   END_IF;
   "CV60PosInit" := #_w7;
   IF #_w7 THEN "PLC_to_Epics".CV60.sSetVAuto := 0.0; END_IF;
   #_w8 := #_w2 AND NOT "CV61_ManAuto";
   IF #_w8 THEN
       "unscal_ret_val_7" := UNSCALE(in := 0.0,
                               hi_lim := 100.0,
                               lo_lim := 0.0,
                               bipolar := "always_0",
                               out => "CMD_CV_61");
   END_IF;
   "CV61PosInit" := #_w8;
   IF #_w8 THEN "PLC_to_Epics".CV61.sSetVAuto := 0.0; END_IF;
   IF #_w2 THEN
       "unscal_ret_val_asco_2" := UNSCALE(in := 100.0,
                               hi_lim := 100.0,
                               lo_lim := 0.0,
                               bipolar := "always_0",
                               out => "Sana_ASCO_2");
   END_IF;
   "ASCO2PosInit" := #_w2;
   IF #_w2 THEN
       "ReguleCV61ON" := FALSE;
       "Separators_empty" := FALSE;
   END_IF;
END_REGION

REGION Network 12: Vanne En Position Initial
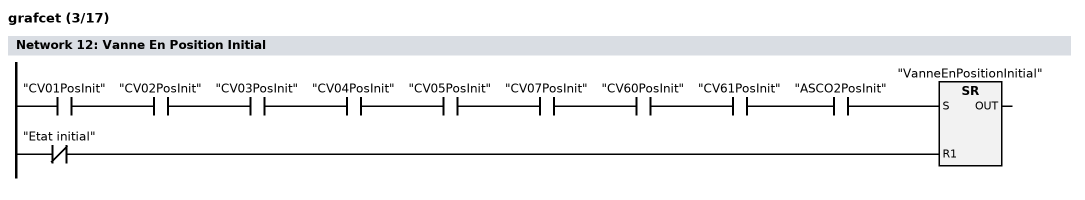
   RUNG wire#powerrail
      Contact( "CV01PosInit" )
      Contact( "CV02PosInit" )
      Contact( "CV03PosInit" )
      Contact( "CV04PosInit" )
      Contact( "CV05PosInit" )
      Contact( "CV07PosInit" )
      Contact( "CV60PosInit" )
      Contact( "CV61PosInit" )
      Contact( "ASCO2PosInit" )
      S_SR(operand := "VanneEnPositionInitial", r1 := wire#w1)
   END_RUNG
   RUNG wire#powerrail
      I_Contact( "Etat initial" )
   END_RUNG wire#w1
   // the same network as SCL:
   IF "CV01PosInit" AND "CV02PosInit" AND "CV03PosInit" AND "CV04PosInit" AND "CV05PosInit" AND "CV07PosInit" AND "CV60PosInit" AND "CV61PosInit" AND "ASCO2PosInit" THEN
       "VanneEnPositionInitial" := TRUE;   // SR flip-flop
   END_IF;
   IF NOT "Etat initial" THEN "VanneEnPositionInitial" := FALSE; END_IF;
END_REGION

REGION Network 13: config vanne etat conditionnement
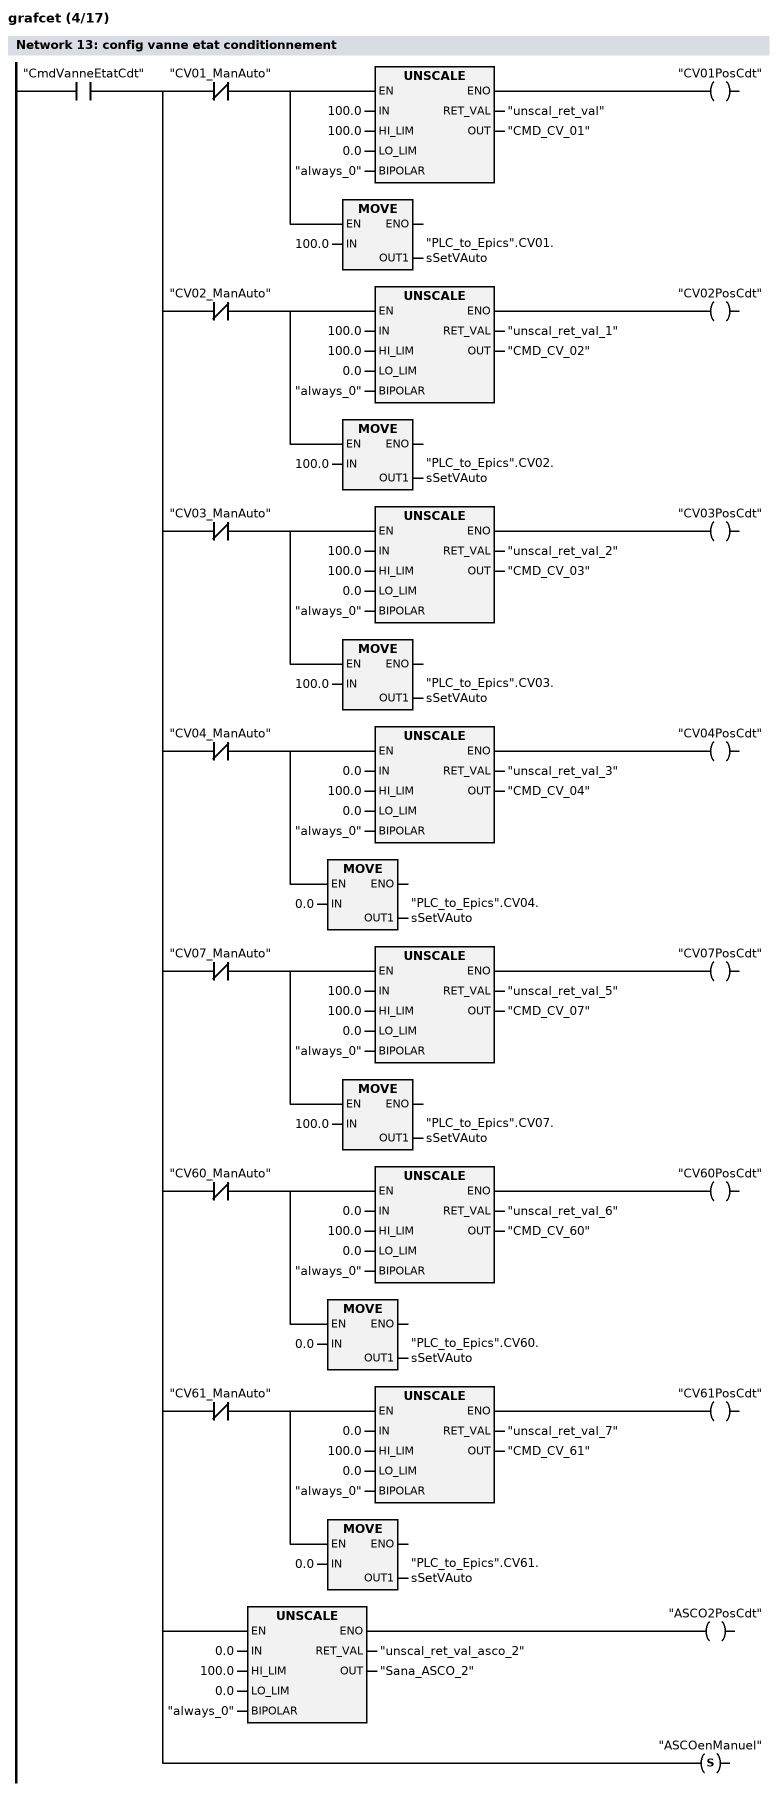
   // ENO of a box is taken as its EN; it also drops when the box reports an error
   #_w1 := "CmdVanneEtatCdt" AND NOT "CV01_ManAuto";
   #_w2 := "CmdVanneEtatCdt";
   IF #_w1 THEN
       "unscal_ret_val" := UNSCALE(IN := 100.0,
                               HI_LIM := 100.0,
                               LO_LIM := 0.0,
                               BIPOLAR := "always_0",
                               OUT => "CMD_CV_01");
   END_IF;
   "CV01PosCdt" := #_w1;
   IF #_w1 THEN "PLC_to_Epics".CV01.sSetVAuto := 100.0; END_IF;
   #_w3 := #_w2 AND NOT "CV02_ManAuto";
   IF #_w3 THEN
       "unscal_ret_val_1" := UNSCALE(IN := 100.0,
                               HI_LIM := 100.0,
                               LO_LIM := 0.0,
                               BIPOLAR := "always_0",
                               OUT => "CMD_CV_02");
   END_IF;
   "CV02PosCdt" := #_w3;
   IF #_w3 THEN "PLC_to_Epics".CV02.sSetVAuto := 100.0; END_IF;
   #_w4 := #_w2 AND NOT "CV03_ManAuto";
   IF #_w4 THEN
       "unscal_ret_val_2" := UNSCALE(IN := 100.0,
                               HI_LIM := 100.0,
                               LO_LIM := 0.0,
                               BIPOLAR := "always_0",
                               OUT => "CMD_CV_03");
   END_IF;
   "CV03PosCdt" := #_w4;
   IF #_w4 THEN "PLC_to_Epics".CV03.sSetVAuto := 100.0; END_IF;
   #_w5 := #_w2 AND NOT "CV04_ManAuto";
   IF #_w5 THEN
       "unscal_ret_val_3" := UNSCALE(IN := 0.0,
                               HI_LIM := 100.0,
                               LO_LIM := 0.0,
                               BIPOLAR := "always_0",
                               OUT => "CMD_CV_04");
   END_IF;
   "CV04PosCdt" := #_w5;
   IF #_w5 THEN "PLC_to_Epics".CV04.sSetVAuto := 0.0; END_IF;
   #_w6 := #_w2 AND NOT "CV07_ManAuto";
   IF #_w6 THEN
       "unscal_ret_val_5" := UNSCALE(IN := 100.0,
                               HI_LIM := 100.0,
                               LO_LIM := 0.0,
                               BIPOLAR := "always_0",
                               OUT => "CMD_CV_07");
   END_IF;
   "CV07PosCdt" := #_w6;
   IF #_w6 THEN "PLC_to_Epics".CV07.sSetVAuto := 100.0; END_IF;
   #_w7 := #_w2 AND NOT "CV60_ManAuto";
   IF #_w7 THEN
       "unscal_ret_val_6" := UNSCALE(IN := 0.0,
                               HI_LIM := 100.0,
                               LO_LIM := 0.0,
                               BIPOLAR := "always_0",
                               OUT => "CMD_CV_60");
   END_IF;
   "CV60PosCdt" := #_w7;
   IF #_w7 THEN "PLC_to_Epics".CV60.sSetVAuto := 0.0; END_IF;
   #_w8 := #_w2 AND NOT "CV61_ManAuto";
   IF #_w8 THEN
       "unscal_ret_val_7" := UNSCALE(IN := 0.0,
                               HI_LIM := 100.0,
                               LO_LIM := 0.0,
                               BIPOLAR := "always_0",
                               OUT => "CMD_CV_61");
   END_IF;
   "CV61PosCdt" := #_w8;
   IF #_w8 THEN "PLC_to_Epics".CV61.sSetVAuto := 0.0; END_IF;
   IF #_w2 THEN
       "unscal_ret_val_asco_2" := UNSCALE(IN := 0.0,
                               HI_LIM := 100.0,
                               LO_LIM := 0.0,
                               BIPOLAR := "always_0",
                               OUT => "Sana_ASCO_2");
   END_IF;
   "ASCO2PosCdt" := #_w2;
   IF #_w2 THEN "ASCOenManuel" := TRUE; END_IF;
END_REGION

REGION Network 14: Vanne En Position Cdt
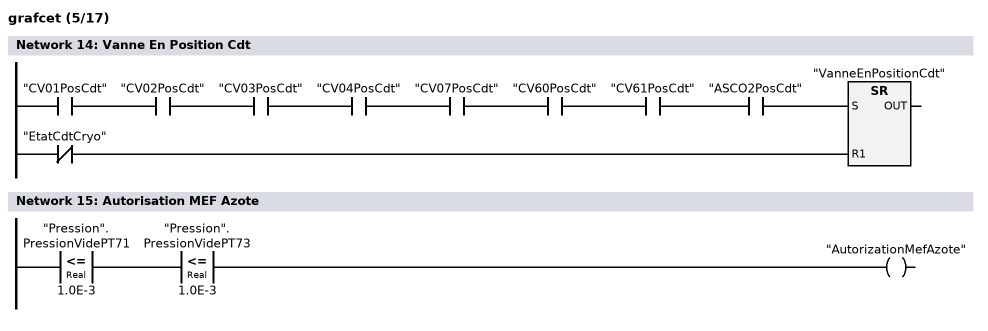
   RUNG wire#powerrail
      Contact( "CV01PosCdt" )
      Contact( "CV02PosCdt" )
      Contact( "CV03PosCdt" )
      Contact( "CV04PosCdt" )
      Contact( "CV07PosCdt" )
      Contact( "CV60PosCdt" )
      Contact( "CV61PosCdt" )
      Contact( "ASCO2PosCdt" )
      S_SR(operand := "VanneEnPositionCdt", r1 := wire#w1)
   END_RUNG
   RUNG wire#powerrail
      I_Contact( "EtatCdtCryo" )
   END_RUNG wire#w1
   // the same network as SCL:
   IF "CV01PosCdt" AND "CV02PosCdt" AND "CV03PosCdt" AND "CV04PosCdt" AND "CV07PosCdt" AND "CV60PosCdt" AND "CV61PosCdt" AND "ASCO2PosCdt" THEN
       "VanneEnPositionCdt" := TRUE;   // SR flip-flop
   END_IF;
   IF NOT "EtatCdtCryo" THEN "VanneEnPositionCdt" := FALSE; END_IF;
END_REGION

REGION Network 15: Autorisation MEF Azote
   RUNG wire#powerrail
      { S7_Templates := "SrcType := Real" } LE_Contact(in1 := "Pression".PressionVidePT71, in2 := 1.0E-3)
      { S7_Templates := "SrcType := Real" } LE_Contact(in1 := "Pression".PressionVidePT73, in2 := 1.0E-3)
      Coil( "AutorizationMefAzote" )
   END_RUNG
   // the same network as SCL:
   "AutorizationMefAzote" := ("Pression".PressionVidePT71 <= 1.0E-3) AND ("Pression".PressionVidePT73 <= 1.0E-3);
END_REGION

REGION Network 16: config vannes init mode & regule cv61 on
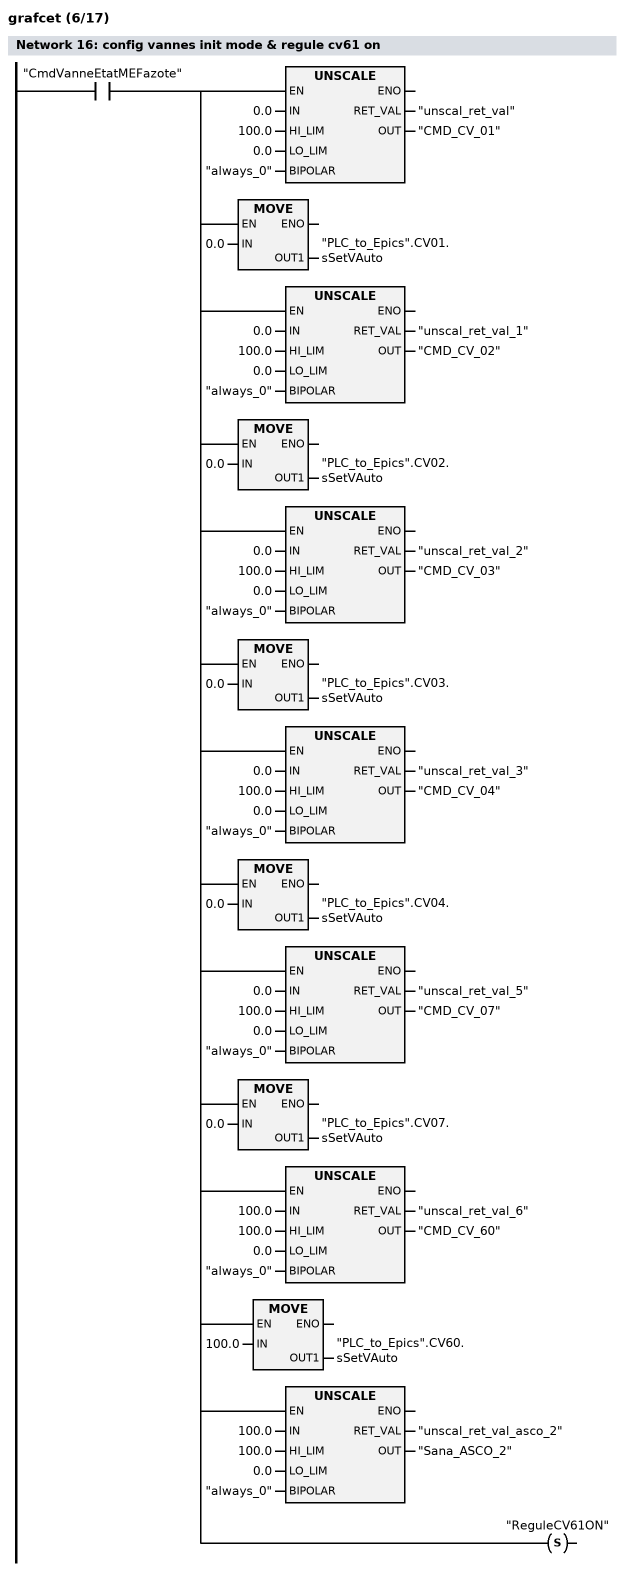
   #_w1 := "CmdVanneEtatMEFazote";
   IF #_w1 THEN
       "unscal_ret_val" := UNSCALE(in := 0.0,
                               hi_lim := 100.0,
                               lo_lim := 0.0,
                               bipolar := "always_0",
                               out => "CMD_CV_01");
       "PLC_to_Epics".CV01.sSetVAuto := 0.0;
       "unscal_ret_val_1" := UNSCALE(in := 0.0,
                               hi_lim := 100.0,
                               lo_lim := 0.0,
                               bipolar := "always_0",
                               out => "CMD_CV_02");
       "PLC_to_Epics".CV02.sSetVAuto := 0.0;
       "unscal_ret_val_2" := UNSCALE(in := 0.0,
                               hi_lim := 100.0,
                               lo_lim := 0.0,
                               bipolar := "always_0",
                               out => "CMD_CV_03");
       "PLC_to_Epics".CV03.sSetVAuto := 0.0;
       "unscal_ret_val_3" := UNSCALE(in := 0.0,
                               hi_lim := 100.0,
                               lo_lim := 0.0,
                               bipolar := "always_0",
                               out => "CMD_CV_04");
       "PLC_to_Epics".CV04.sSetVAuto := 0.0;
       "unscal_ret_val_5" := UNSCALE(in := 0.0,
                               hi_lim := 100.0,
                               lo_lim := 0.0,
                               bipolar := "always_0",
                               out => "CMD_CV_07");
       "PLC_to_Epics".CV07.sSetVAuto := 0.0;
       "unscal_ret_val_6" := UNSCALE(in := 100.0,
                               hi_lim := 100.0,
                               lo_lim := 0.0,
                               bipolar := "always_0",
                               out => "CMD_CV_60");
       "PLC_to_Epics".CV60.sSetVAuto := 100.0;
       "unscal_ret_val_asco_2" := UNSCALE(in := 100.0,
                               hi_lim := 100.0,
                               lo_lim := 0.0,
                               bipolar := "always_0",
                               out => "Sana_ASCO_2");
       "ReguleCV61ON" := TRUE;
   END_IF;
END_REGION

REGION Network 17: Régule CV61 seuil (desactive)
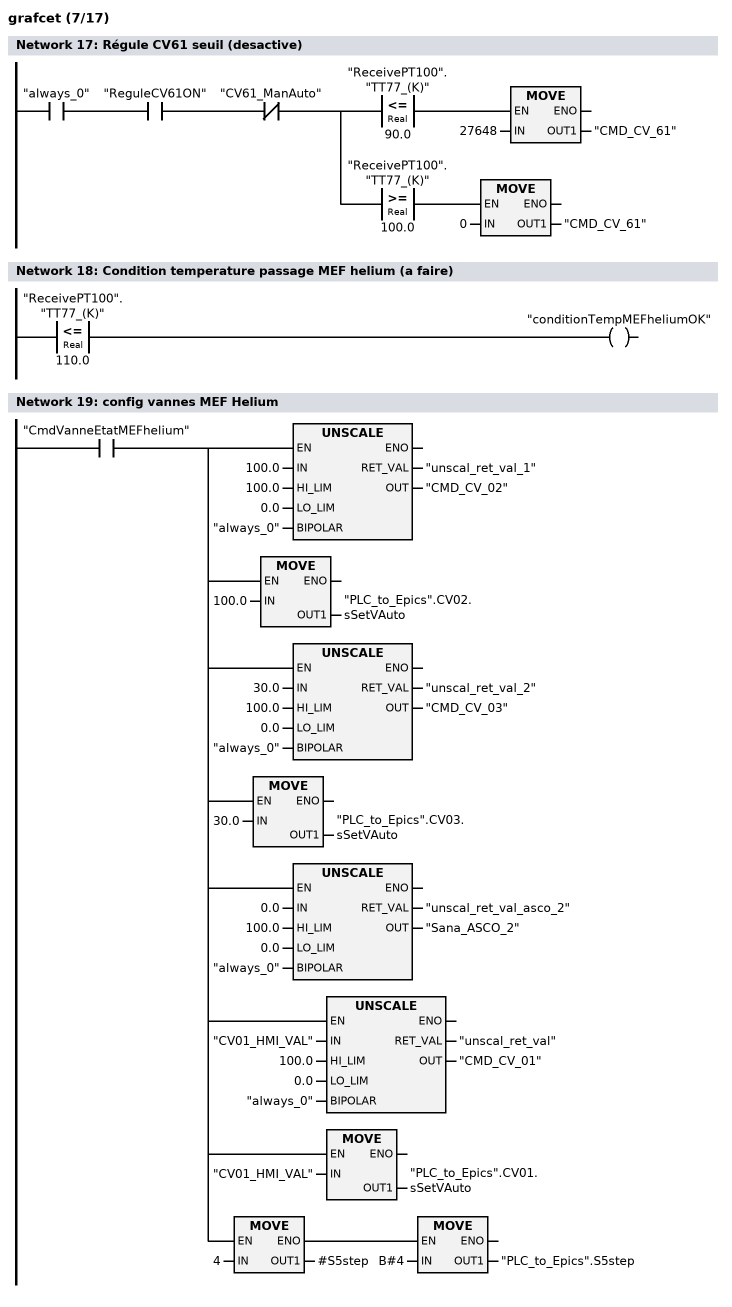
   RUNG wire#powerrail
      Contact( "always_0" )
      Contact( "ReguleCV61ON" )
      I_Contact( "CV61_ManAuto" )
      wire#w1
      { S7_Templates := "SrcType := Real" } LE_Contact(in1 := "ReceivePT100"."TT77_(K)", in2 := 90.0)
      { S7_GenerateENO := "TRUE" } Move(in := 27648, out1 => "CMD_CV_61")
   END_RUNG
   RUNG wire#w1
      { S7_Templates := "SrcType := Real" } GE_Contact(in1 := "ReceivePT100"."TT77_(K)", in2 := 100.0)
      { S7_GenerateENO := "TRUE" } Move(in := 0, out1 => "CMD_CV_61")
   END_RUNG
   // the same network as SCL:
   #_w1 := "always_0" AND "ReguleCV61ON" AND NOT "CV61_ManAuto";
   IF #_w1 AND ("ReceivePT100"."TT77_(K)" <= 90.0) THEN "CMD_CV_61" := 27648; END_IF;
   IF #_w1 AND ("ReceivePT100"."TT77_(K)" >= 100.0) THEN "CMD_CV_61" := 0; END_IF;
END_REGION

REGION Network 18: Condition temperature passage MEF helium (a faire)
   RUNG wire#powerrail
      { S7_Templates := "SrcType := Real" } LE_Contact(in1 := "ReceivePT100"."TT77_(K)", in2 := 110.0)
      Coil( "conditionTempMEFheliumOK" )
   END_RUNG
   // the same network as SCL:
   "conditionTempMEFheliumOK" := "ReceivePT100"."TT77_(K)" <= 110.0;
END_REGION

REGION Network 19: config vannes MEF Helium
   // ENO of a box is taken as its EN; it also drops when the box reports an error
   #_w1 := "CmdVanneEtatMEFhelium";
   IF #_w1 THEN
       "unscal_ret_val_1" := UNSCALE(IN := 100.0,
                               HI_LIM := 100.0,
                               LO_LIM := 0.0,
                               BIPOLAR := "always_0",
                               OUT => "CMD_CV_02");
       "PLC_to_Epics".CV02.sSetVAuto := 100.0;
       "unscal_ret_val_2" := UNSCALE(IN := 30.0,
                               HI_LIM := 100.0,
                               LO_LIM := 0.0,
                               BIPOLAR := "always_0",
                               OUT => "CMD_CV_03");
       "PLC_to_Epics".CV03.sSetVAuto := 30.0;
       "unscal_ret_val_asco_2" := UNSCALE(IN := 0.0,
                               HI_LIM := 100.0,
                               LO_LIM := 0.0,
                               BIPOLAR := "always_0",
                               OUT => "Sana_ASCO_2");
       "unscal_ret_val" := UNSCALE(IN := "CV01_HMI_VAL",
                               HI_LIM := 100.0,
                               LO_LIM := 0.0,
                               BIPOLAR := "always_0",
                               OUT => "CMD_CV_01");
       "PLC_to_Epics".CV01.sSetVAuto := "CV01_HMI_VAL";
       #S5step := 4;
       "PLC_to_Epics".S5step := B#4;
   END_IF;
END_REGION

REGION Network 20: LHe cooling down - Set step 6 (maybe setting CV03 is not needed here (done in the next network)!!!!!
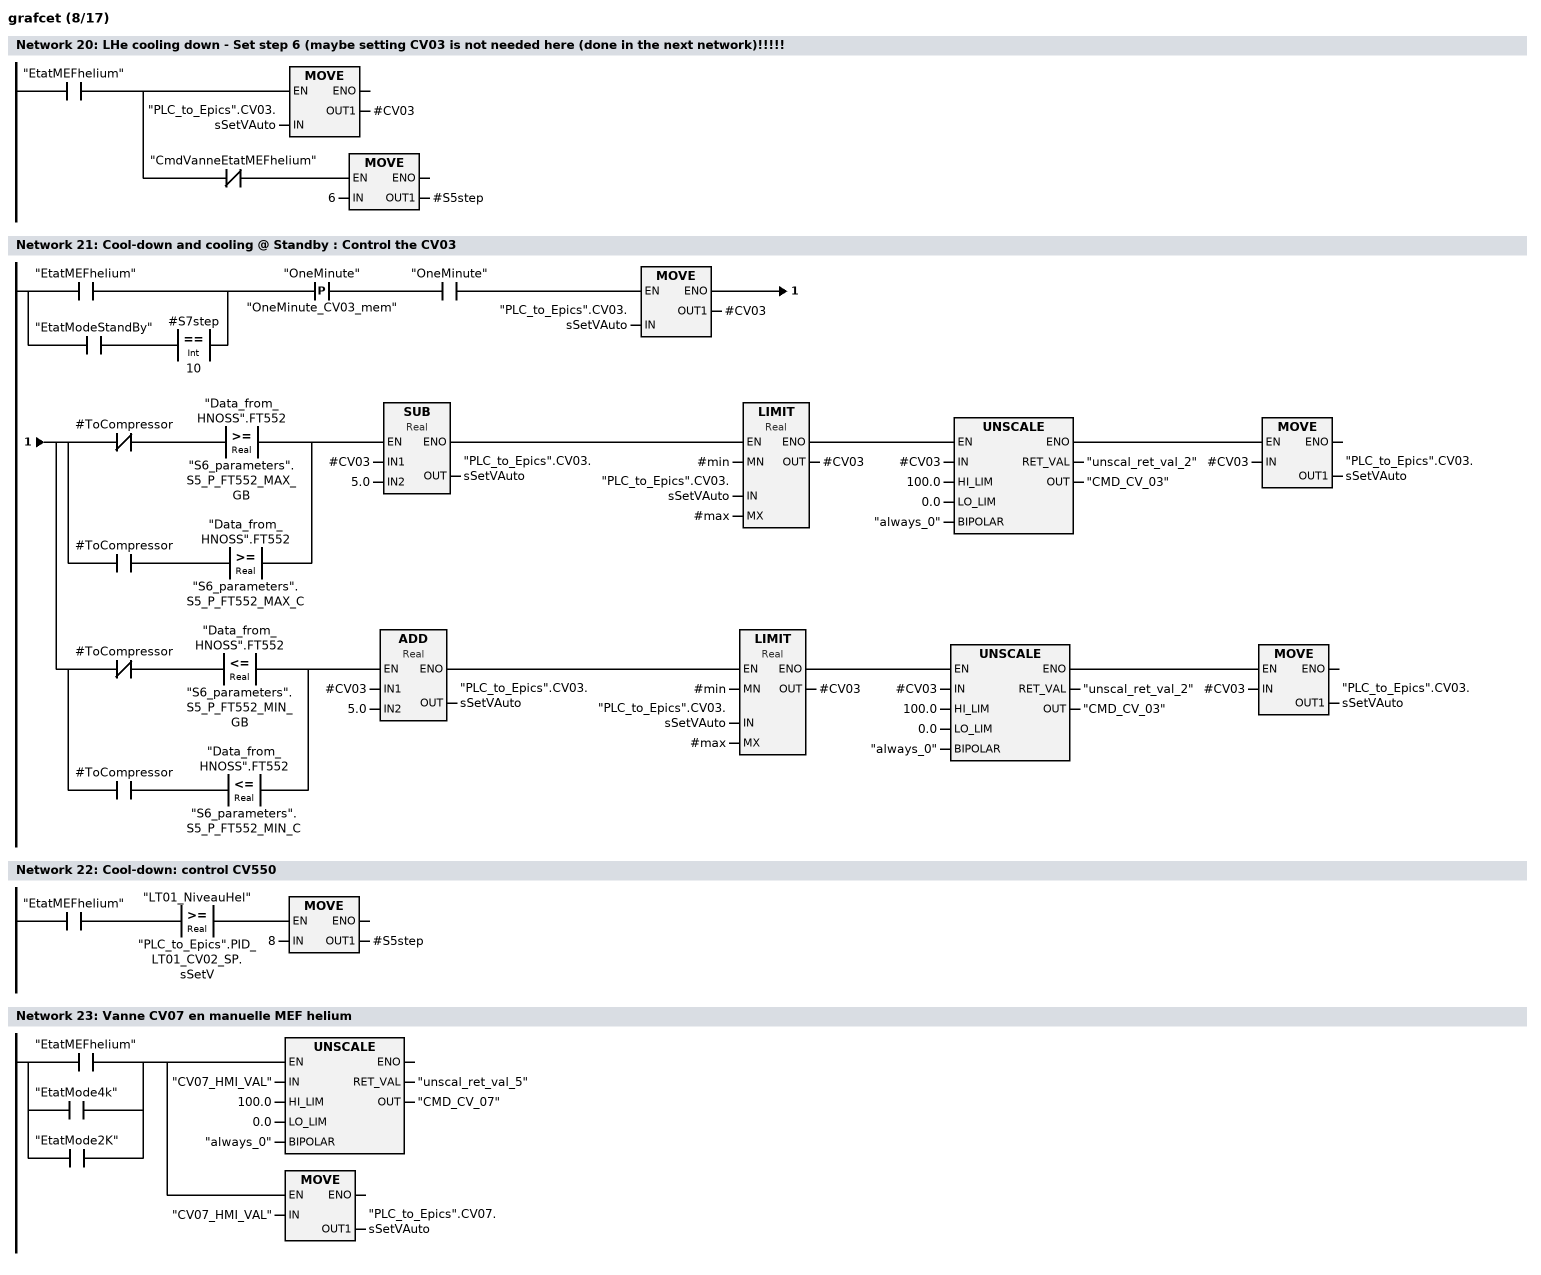
   RUNG wire#powerrail
      Contact( "EtatMEFhelium" )
      wire#w1
      { S7_GenerateENO := "TRUE" } Move(in := "PLC_to_Epics".CV03.sSetVAuto, out1 => #CV03)
   END_RUNG
   RUNG wire#w1
      I_Contact( "CmdVanneEtatMEFhelium" )
      { S7_GenerateENO := "TRUE" } Move(in := 6, out1 => #S5step)
   END_RUNG
   // the same network as SCL:
   IF "EtatMEFhelium" THEN #CV03 := "PLC_to_Epics".CV03.sSetVAuto; END_IF;
   IF "EtatMEFhelium" AND NOT "CmdVanneEtatMEFhelium" THEN #S5step := 6; END_IF;
END_REGION

REGION Network 21: Cool-down and cooling @ Standby : Control the CV03
   // ENO of a box is taken as its EN; it also drops when the box reports an error
   #_w1 := ("EtatMEFhelium" OR ("EtatModeStandBy" AND (#S7step = 10))) AND "OneMinute" AND NOT "OneMinute_CV03_mem";   // rising edge of "OneMinute"
   "OneMinute_CV03_mem" := "OneMinute";
   #_w2 := #_w1 AND "OneMinute";
   IF #_w2 THEN #CV03 := "PLC_to_Epics".CV03.sSetVAuto; END_IF;
   IF #_w2 AND ((NOT #ToCompressor AND ("Data_from_HNOSS".FT552 >= "S6_parameters".S5_P_FT552_MAX_GB)) OR (#ToCompressor AND ("Data_from_HNOSS".FT552 >= "S6_parameters".S5_P_FT552_MAX_C))) THEN
       "PLC_to_Epics".CV03.sSetVAuto := #CV03 - 5.0;
       #CV03 := LIMIT(MN := #min, IN := "PLC_to_Epics".CV03.sSetVAuto, MX := #max);
   END_IF;
   #_w3 := #_w2 AND ((NOT #ToCompressor AND ("Data_from_HNOSS".FT552 >= "S6_parameters".S5_P_FT552_MAX_GB)) OR (#ToCompressor AND ("Data_from_HNOSS".FT552 >= "S6_parameters".S5_P_FT552_MAX_C)));
   IF #_w3 THEN
       "unscal_ret_val_2" := UNSCALE(IN := #CV03,
                               HI_LIM := 100.0,
                               LO_LIM := 0.0,
                               BIPOLAR := "always_0",
                               OUT => "CMD_CV_03");
       "PLC_to_Epics".CV03.sSetVAuto := #CV03;
   END_IF;
   IF #_w2 AND ((NOT #ToCompressor AND ("Data_from_HNOSS".FT552 <= "S6_parameters".S5_P_FT552_MIN_GB)) OR (#ToCompressor AND ("Data_from_HNOSS".FT552 <= "S6_parameters".S5_P_FT552_MIN_C))) THEN
       "PLC_to_Epics".CV03.sSetVAuto := #CV03 + 5.0;
       #CV03 := LIMIT(MN := #min, IN := "PLC_to_Epics".CV03.sSetVAuto, MX := #max);
   END_IF;
   #_w4 := #_w2 AND ((NOT #ToCompressor AND ("Data_from_HNOSS".FT552 <= "S6_parameters".S5_P_FT552_MIN_GB)) OR (#ToCompressor AND ("Data_from_HNOSS".FT552 <= "S6_parameters".S5_P_FT552_MIN_C)));
   IF #_w4 THEN
       "unscal_ret_val_2" := UNSCALE(IN := #CV03,
                               HI_LIM := 100.0,
                               LO_LIM := 0.0,
                               BIPOLAR := "always_0",
                               OUT => "CMD_CV_03");
       "PLC_to_Epics".CV03.sSetVAuto := #CV03;
   END_IF;
END_REGION

REGION Network 22: Cool-down: control CV550
   RUNG wire#powerrail
      Contact( "EtatMEFhelium" )
      { S7_Templates := "SrcType := Real" } GE_Contact(in1 := "LT01_NiveauHel", in2 := "PLC_to_Epics".PID_LT01_CV02_SP.sSetV)
      { S7_GenerateENO := "TRUE" } Move(in := 8, out1 => #S5step)
   END_RUNG
   // the same network as SCL:
   IF "EtatMEFhelium" AND ("LT01_NiveauHel" >= "PLC_to_Epics".PID_LT01_CV02_SP.sSetV) THEN
       #S5step := 8;
   END_IF;
END_REGION

REGION Network 23: Vanne CV07 en manuelle MEF helium
   #_w1 := "EtatMEFhelium" OR "EtatMode4k" OR "EtatMode2K";
   IF #_w1 THEN
       "unscal_ret_val_5" := UNSCALE(in := "CV07_HMI_VAL",
                               hi_lim := 100.0,
                               lo_lim := 0.0,
                               bipolar := "always_0",
                               out => "CMD_CV_07");
       "PLC_to_Epics".CV07.sSetVAuto := "CV07_HMI_VAL";
   END_IF;
END_REGION

REGION Network 24: Vanne CV01 en manuelle MEF helium
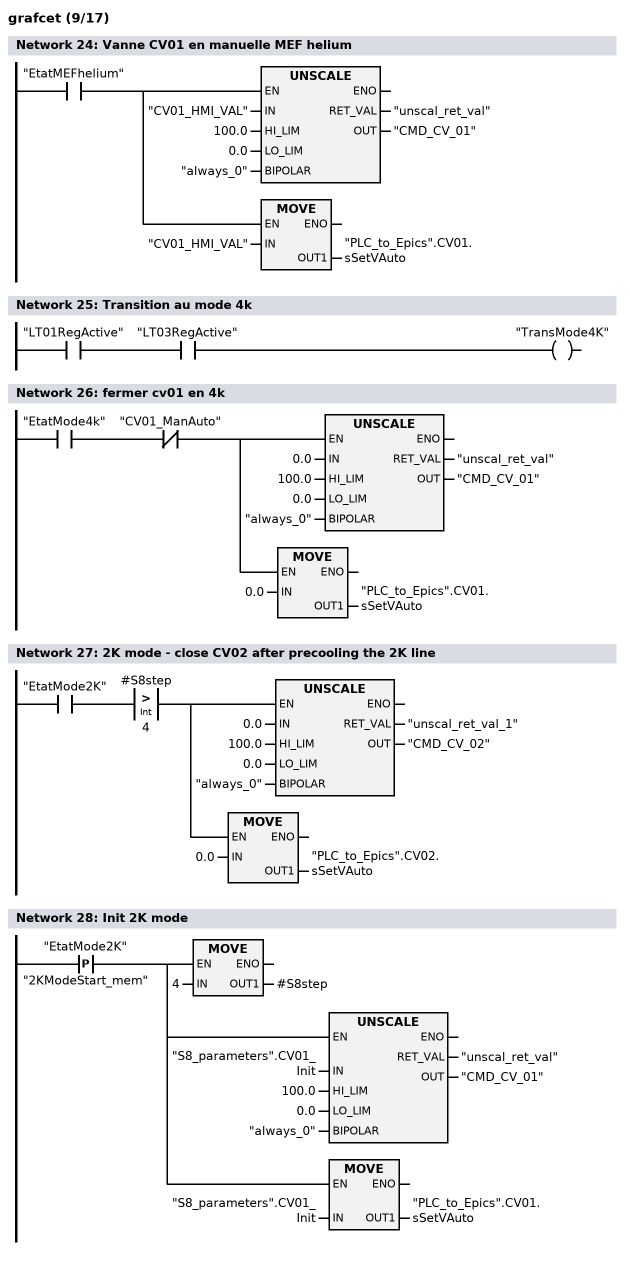
   #_w1 := "EtatMEFhelium";
   IF #_w1 THEN
       "unscal_ret_val" := UNSCALE(in := "CV01_HMI_VAL",
                               hi_lim := 100.0,
                               lo_lim := 0.0,
                               bipolar := "always_0",
                               out => "CMD_CV_01");
       "PLC_to_Epics".CV01.sSetVAuto := "CV01_HMI_VAL";
   END_IF;
END_REGION

REGION Network 25: Transition au mode 4k
   RUNG wire#powerrail
      Contact( "LT01RegActive" )
      Contact( "LT03RegActive" )
      Coil( "TransMode4K" )
   END_RUNG
   // the same network as SCL:
   "TransMode4K" := "LT01RegActive" AND "LT03RegActive";
END_REGION

REGION Network 26: fermer cv01 en 4k
   #_w1 := "EtatMode4k" AND NOT "CV01_ManAuto";
   IF #_w1 THEN
       "unscal_ret_val" := UNSCALE(in := 0.0,
                               hi_lim := 100.0,
                               lo_lim := 0.0,
                               bipolar := "always_0",
                               out => "CMD_CV_01");
       "PLC_to_Epics".CV01.sSetVAuto := 0.0;
   END_IF;
END_REGION

REGION Network 27: 2K mode - close CV02 after precooling the 2K line
   #_w1 := "EtatMode2K" AND (#S8step > 4);
   IF #_w1 THEN
       "unscal_ret_val_1" := UNSCALE(IN := 0.0,
                               HI_LIM := 100.0,
                               LO_LIM := 0.0,
                               BIPOLAR := "always_0",
                               OUT => "CMD_CV_02");
       "PLC_to_Epics".CV02.sSetVAuto := 0.0;
   END_IF;
END_REGION

REGION Network 28: Init 2K mode
   #_w1 := "EtatMode2K" AND NOT "2KModeStart_mem";   // rising edge of "EtatMode2K"
   "2KModeStart_mem" := "EtatMode2K";
   IF #_w1 THEN
       #S8step := 4;
       "unscal_ret_val" := UNSCALE(IN := "S8_parameters".CV01_Init,
                               HI_LIM := 100.0,
                               LO_LIM := 0.0,
                               BIPOLAR := "always_0",
                               OUT => "CMD_CV_01");
       "PLC_to_Epics".CV01.sSetVAuto := "S8_parameters".CV01_Init;
   END_IF;
END_REGION

REGION Network 29: 2K mode - precooling (step4)
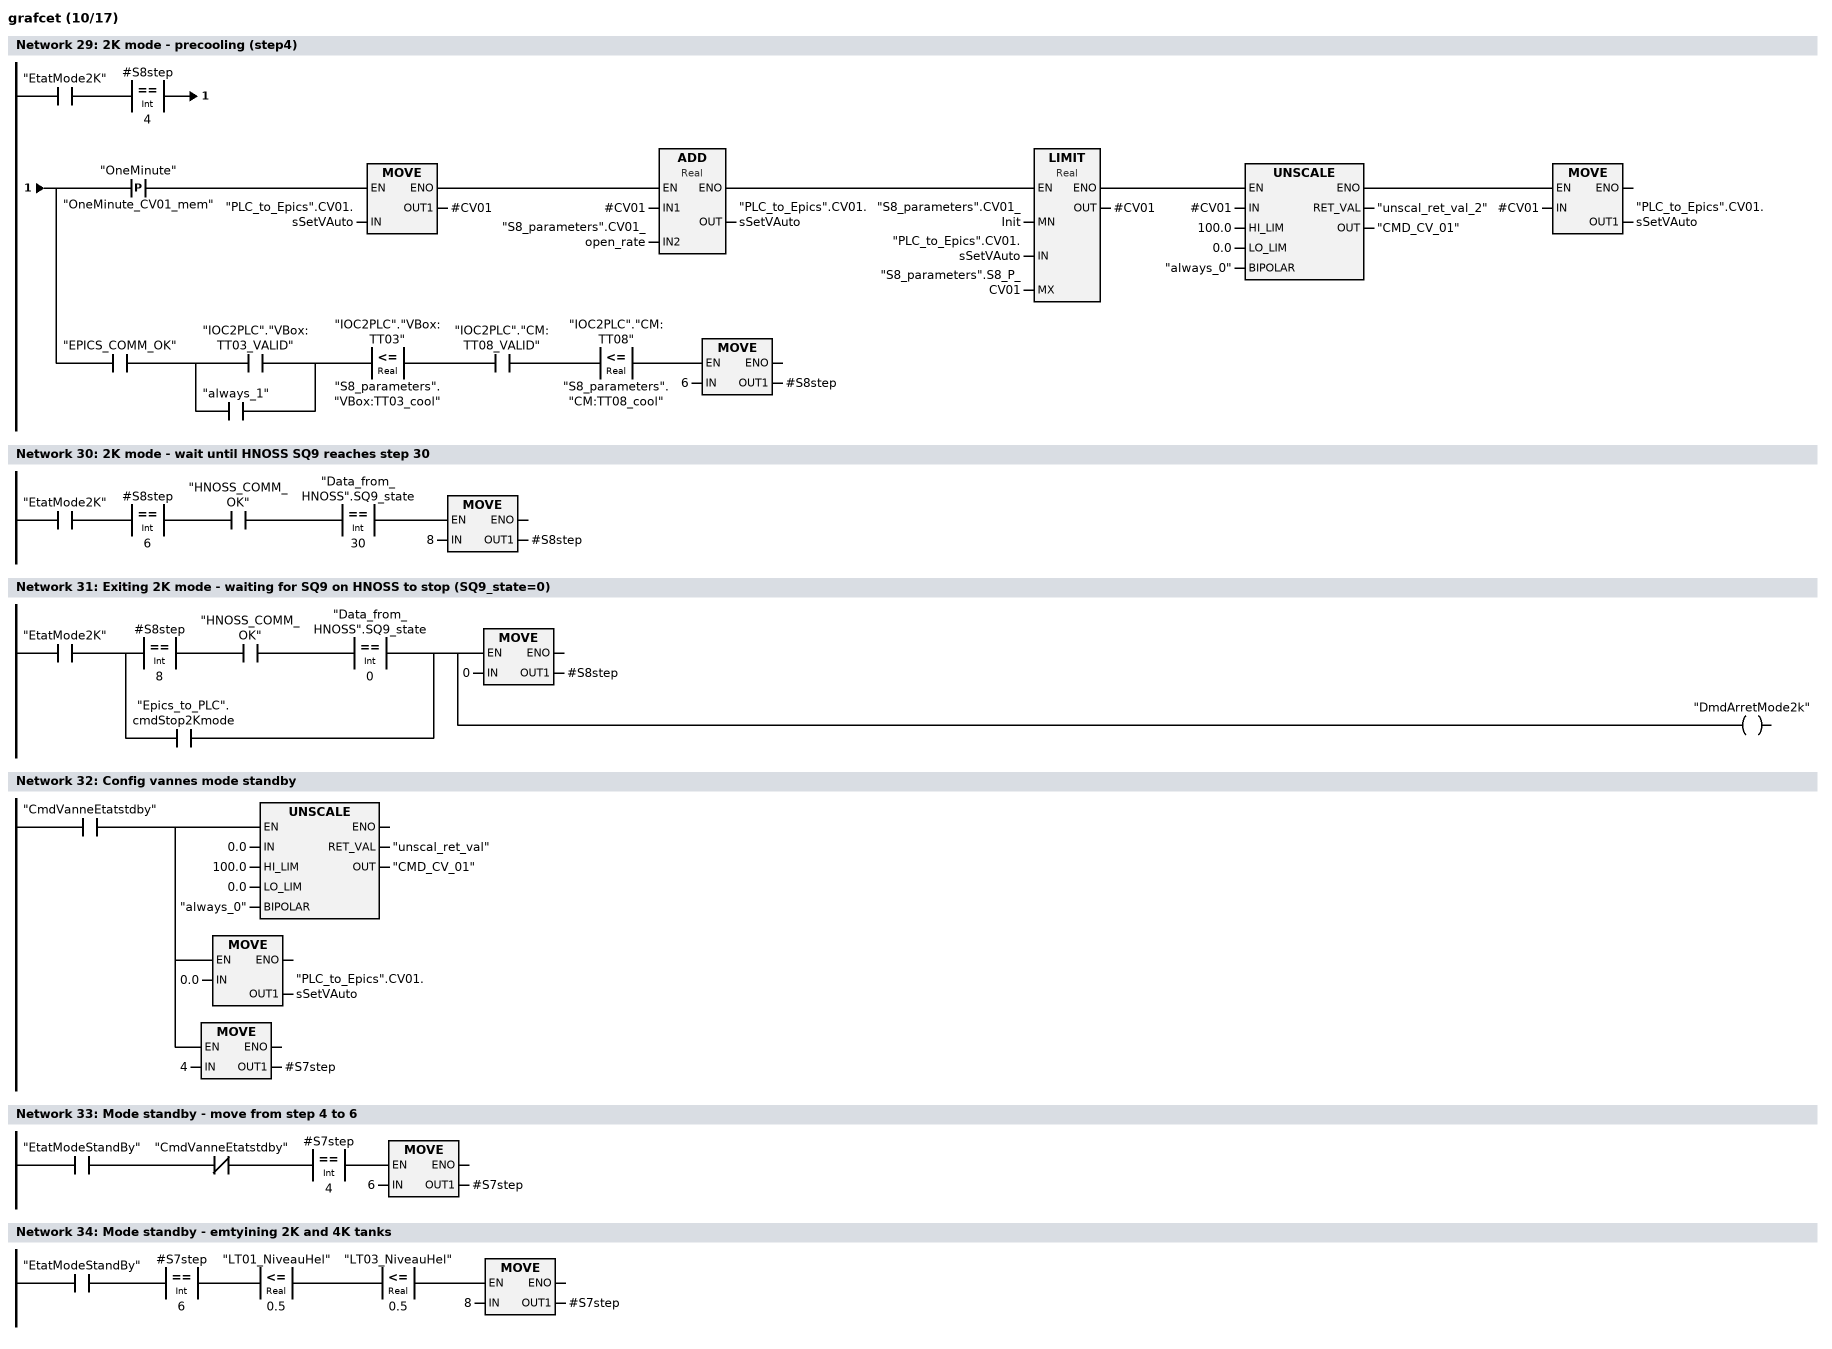
   // ENO of a box is taken as its EN; it also drops when the box reports an error
   #_w1 := "EtatMode2K" AND (#S8step = 4);
   #_w2 := #_w1 AND "OneMinute" AND NOT "OneMinute_CV01_mem";   // rising edge of "OneMinute"
   "OneMinute_CV01_mem" := "OneMinute";
   IF #_w2 THEN
       #CV01 := "PLC_to_Epics".CV01.sSetVAuto;
       "PLC_to_Epics".CV01.sSetVAuto := #CV01 + "S8_parameters".CV01_open_rate;
       #CV01 := LIMIT(MN := "S8_parameters".CV01_Init, IN := "PLC_to_Epics".CV01.sSetVAuto, MX := "S8_parameters".S8_P_CV01);
       "unscal_ret_val_2" := UNSCALE(IN := #CV01,
                               HI_LIM := 100.0,
                               LO_LIM := 0.0,
                               BIPOLAR := "always_0",
                               OUT => "CMD_CV_01");
       "PLC_to_Epics".CV01.sSetVAuto := #CV01;
   END_IF;
   IF #_w1 AND "EPICS_COMM_OK" AND ("IOC2PLC"."VBox:TT03_VALID" OR "always_1") AND ("IOC2PLC"."VBox:TT03" <= "S8_parameters"."VBox:TT03_cool") AND "IOC2PLC"."CM:TT08_VALID" AND ("IOC2PLC"."CM:TT08" <= "S8_parameters"."CM:TT08_cool") THEN
       #S8step := 6;
   END_IF;
END_REGION

REGION Network 30: 2K mode - wait until HNOSS SQ9 reaches step 30
   RUNG wire#powerrail
      Contact( "EtatMode2K" )
      { S7_Templates := "SrcType := Int" } EQ_Contact(in1 := #S8step, in2 := 6)
      Contact( "HNOSS_COMM_OK" )
      { S7_Templates := "SrcType := Int" } EQ_Contact(in1 := "Data_from_HNOSS".SQ9_state, in2 := 30)
      { S7_GenerateENO := "TRUE" } Move(in := 8, out1 => #S8step)
   END_RUNG
   // the same network as SCL:
   IF "EtatMode2K" AND (#S8step = 6) AND "HNOSS_COMM_OK" AND ("Data_from_HNOSS".SQ9_state = 30) THEN
       #S8step := 8;
   END_IF;
END_REGION

REGION Network 31: Exiting 2K mode - waiting for SQ9 on HNOSS to stop (SQ9_state=0)
   RUNG wire#powerrail
      Contact( "EtatMode2K" )
      wire#w1
      { S7_Templates := "SrcType := Int" } EQ_Contact(in1 := #S8step, in2 := 8)
      Contact( "HNOSS_COMM_OK" )
      { S7_Templates := "SrcType := Int" } EQ_Contact(in1 := "Data_from_HNOSS".SQ9_state, in2 := 0)
      wire#w2
      { S7_GenerateENO := "TRUE" } Move(in := 0, out1 => #S8step)
   END_RUNG
   RUNG wire#w1
      Contact( "Epics_to_PLC".cmdStop2Kmode )
   END_RUNG wire#w2
   RUNG wire#w2
      Coil( "DmdArretMode2k" )
   END_RUNG
   // the same network as SCL:
   #_w1 := "EtatMode2K" AND (((#S8step = 8) AND "HNOSS_COMM_OK" AND ("Data_from_HNOSS".SQ9_state = 0)) OR "Epics_to_PLC".cmdStop2Kmode);
   IF #_w1 THEN #S8step := 0; END_IF;
   "DmdArretMode2k" := #_w1;
END_REGION

REGION Network 32: Config vannes mode standby
   #_w1 := "CmdVanneEtatstdby";
   IF #_w1 THEN
       "unscal_ret_val" := UNSCALE(IN := 0.0,
                               HI_LIM := 100.0,
                               LO_LIM := 0.0,
                               BIPOLAR := "always_0",
                               OUT => "CMD_CV_01");
       "PLC_to_Epics".CV01.sSetVAuto := 0.0;
       #S7step := 4;
   END_IF;
END_REGION

REGION Network 33: Mode standby - move from step 4 to 6
   RUNG wire#powerrail
      Contact( "EtatModeStandBy" )
      I_Contact( "CmdVanneEtatstdby" )
      { S7_Templates := "SrcType := Int" } EQ_Contact(in1 := #S7step, in2 := 4)
      { S7_GenerateENO := "TRUE" } Move(in := 6, out1 => #S7step)
   END_RUNG
   // the same network as SCL:
   IF "EtatModeStandBy" AND NOT "CmdVanneEtatstdby" AND (#S7step = 4) THEN #S7step := 6; END_IF;
END_REGION

REGION Network 34: Mode standby - emtyining 2K and 4K tanks
   RUNG wire#powerrail
      Contact( "EtatModeStandBy" )
      { S7_Templates := "SrcType := Int" } EQ_Contact(in1 := #S7step, in2 := 6)
      { S7_Templates := "SrcType := Real" } LE_Contact(in1 := "LT01_NiveauHel", in2 := 0.5)
      { S7_Templates := "SrcType := Real" } LE_Contact(in1 := "LT03_NiveauHel", in2 := 0.5)
      { S7_GenerateENO := "TRUE" } Move(in := 8, out1 => #S7step)
   END_RUNG
   // the same network as SCL:
   IF "EtatModeStandBy" AND (#S7step = 6) AND ("LT01_NiveauHel" <= 0.5) AND ("LT03_NiveauHel" <= 0.5) THEN
       #S7step := 8;
   END_IF;
END_REGION

REGION Network 35: Mode standby - warming up (step8) and cooling (step10)
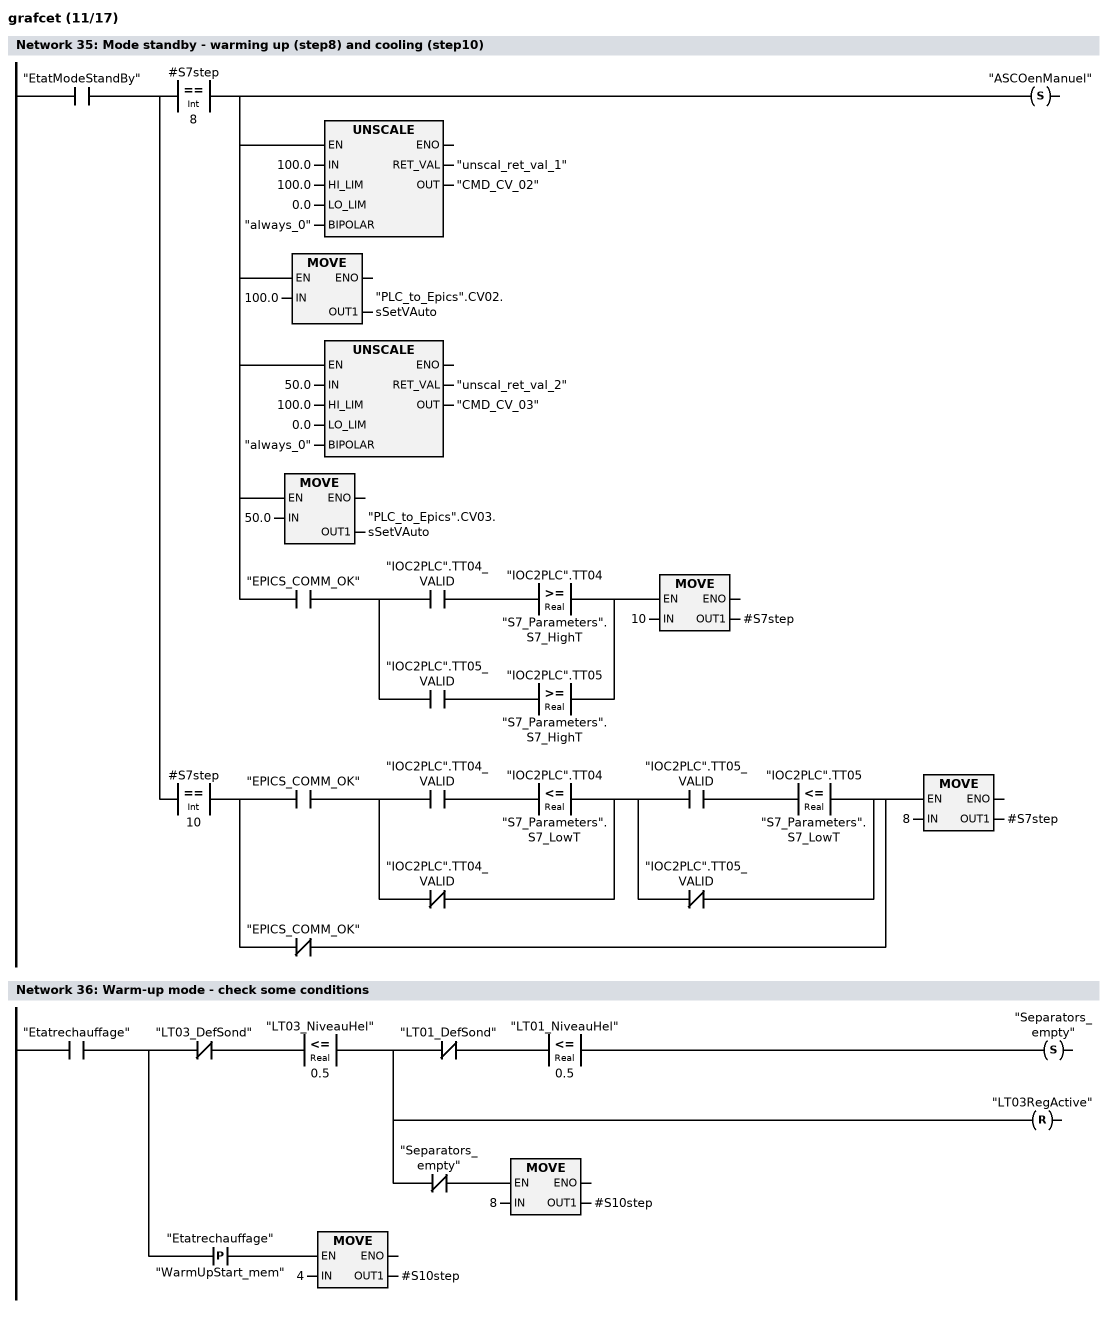
   #_w1 := "EtatModeStandBy" AND (#S7step = 8);
   IF #_w1 THEN "ASCOenManuel" := TRUE; END_IF;
   #_w2 := "EtatModeStandBy";
   IF #_w1 THEN
       "unscal_ret_val_1" := UNSCALE(IN := 100.0,
                               HI_LIM := 100.0,
                               LO_LIM := 0.0,
                               BIPOLAR := "always_0",
                               OUT => "CMD_CV_02");
       "PLC_to_Epics".CV02.sSetVAuto := 100.0;
       "unscal_ret_val_2" := UNSCALE(IN := 50.0,
                               HI_LIM := 100.0,
                               LO_LIM := 0.0,
                               BIPOLAR := "always_0",
                               OUT => "CMD_CV_03");
       "PLC_to_Epics".CV03.sSetVAuto := 50.0;
   END_IF;
   IF #_w1 AND "EPICS_COMM_OK" AND (("IOC2PLC".TT04_VALID AND ("IOC2PLC".TT04 >= "S7_Parameters".S7_HighT)) OR ("IOC2PLC".TT05_VALID AND ("IOC2PLC".TT05 >= "S7_Parameters".S7_HighT))) THEN
       #S7step := 10;
   END_IF;
   IF #_w2 AND (#S7step = 10) AND (("EPICS_COMM_OK" AND (("IOC2PLC".TT04_VALID AND ("IOC2PLC".TT04 <= "S7_Parameters".S7_LowT)) OR NOT "IOC2PLC".TT04_VALID) AND (("IOC2PLC".TT05_VALID AND ("IOC2PLC".TT05 <= "S7_Parameters".S7_LowT)) OR NOT "IOC2PLC".TT05_VALID)) OR NOT "EPICS_COMM_OK") THEN
       #S7step := 8;
   END_IF;
END_REGION

REGION Network 36: Warm-up mode - check some conditions
   RUNG wire#powerrail
      Contact( "Etatrechauffage" )
      wire#w1
      I_Contact( "LT03_DefSond" )
      { S7_Templates := "SrcType := Real" } LE_Contact(in1 := "LT03_NiveauHel", in2 := 0.5)
      wire#w2
      I_Contact( "LT01_DefSond" )
      { S7_Templates := "SrcType := Real" } LE_Contact(in1 := "LT01_NiveauHel", in2 := 0.5)
      S_Coil( "Separators_empty" )
   END_RUNG
   RUNG wire#w2
      R_Coil( "LT03RegActive" )
   END_RUNG
   RUNG wire#w2
      I_Contact( "Separators_empty" )
      { S7_GenerateENO := "TRUE" } Move(in := 8, out1 => #S10step)
   END_RUNG
   RUNG wire#w1
      P_Contact(operand := "Etatrechauffage", bit := "WarmUpStart_mem")
      { S7_GenerateENO := "TRUE" } Move(in := 4, out1 => #S10step)
   END_RUNG
   // the same network as SCL:
   #_w1 := "Etatrechauffage" AND NOT "LT03_DefSond" AND ("LT03_NiveauHel" <= 0.5);
   IF #_w1 AND NOT "LT01_DefSond" AND ("LT01_NiveauHel" <= 0.5) THEN "Separators_empty" := TRUE; END_IF;
   IF #_w1 THEN "LT03RegActive" := FALSE; END_IF;
   IF #_w1 AND NOT "Separators_empty" THEN #S10step := 8; END_IF;
   #_w2 := "Etatrechauffage" AND "Etatrechauffage" AND NOT "WarmUpStart_mem";   // rising edge of "Etatrechauffage"
   "WarmUpStart_mem" := "Etatrechauffage";
   IF #_w2 THEN #S10step := 4; END_IF;
END_REGION

REGION Network 37: Warm-up: set-up the settings of CV01-CV04
   // Set-up the settings depending on the LHe levels in the phase separators
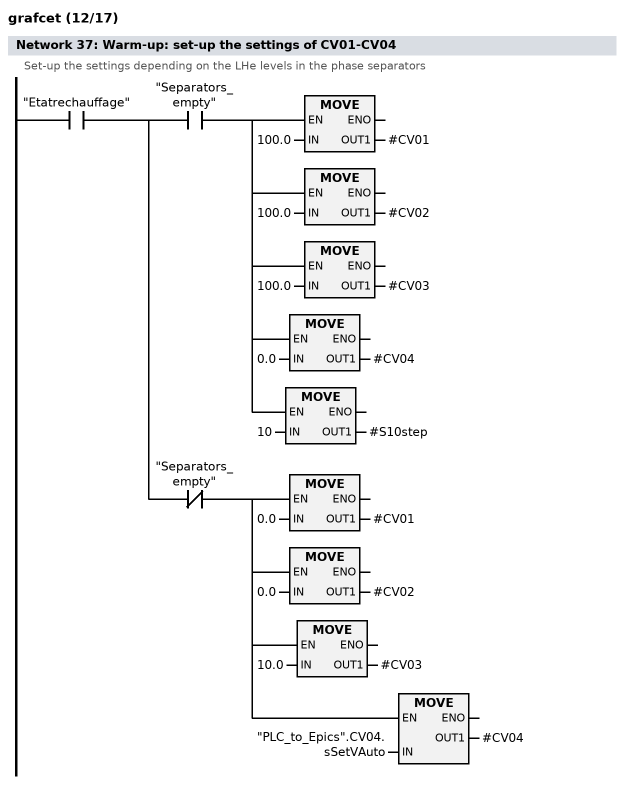
   RUNG wire#powerrail
      Contact( "Etatrechauffage" )
      wire#w1
      Contact( "Separators_empty" )
      wire#w2
      { S7_GenerateENO := "TRUE" } Move(in := 100.0, out1 => #CV01)
   END_RUNG
   RUNG wire#w2
      { S7_GenerateENO := "TRUE" } Move(in := 100.0, out1 => #CV02)
   END_RUNG
   RUNG wire#w2
      { S7_GenerateENO := "TRUE" } Move(in := 100.0, out1 => #CV03)
   END_RUNG
   RUNG wire#w2
      { S7_GenerateENO := "TRUE" } Move(in := 0.0, out1 => #CV04)
   END_RUNG
   RUNG wire#w2
      { S7_GenerateENO := "TRUE" } Move(in := 10, out1 => #S10step)
   END_RUNG
   RUNG wire#w1
      I_Contact( "Separators_empty" )
      wire#w3
      { S7_GenerateENO := "TRUE" } Move(in := 0.0, out1 => #CV01)
   END_RUNG
   RUNG wire#w3
      { S7_GenerateENO := "TRUE" } Move(in := 0.0, out1 => #CV02)
   END_RUNG
   RUNG wire#w3
      { S7_GenerateENO := "TRUE" } Move(in := 10.0, out1 => #CV03)
   END_RUNG
   RUNG wire#w3
      { S7_GenerateENO := "TRUE" } Move(in := "PLC_to_Epics".CV04.sSetVAuto, out1 => #CV04)
   END_RUNG
   // the same network as SCL:
   IF "Etatrechauffage" AND "Separators_empty" THEN
       #CV01 := 100.0;
       #CV02 := 100.0;
       #CV03 := 100.0;
       #CV04 := 0.0;
       #S10step := 10;
   END_IF;
   IF "Etatrechauffage" AND NOT "Separators_empty" THEN
       #CV01 := 0.0;
       #CV02 := 0.0;
       #CV03 := 10.0;
       #CV04 := "PLC_to_Epics".CV04.sSetVAuto;
   END_IF;
END_REGION

REGION Network 38: Mode Rechauffage
   // The heaters are handled in Manage_HEATERS